REGION Network 5
   RUNG wire#powerrail
      { S7_Templates := "SrcType := Int" } EQ_Contact(in1 := #IN0, in2 := 2048)
      { S7_GenerateENO := "TRUE" } Move(in := 4, out1 => #OUT1)
   END_RUNG
   // the same network as SCL:
   IF #IN0 = 2048 THEN #OUT1 := 4; END_IF;
END_REGION

REGION Network 6
   RUNG wire#powerrail
      { S7_Templates := "SrcType := Int" } EQ_Contact(in1 := #IN0, in2 := 4096)
      { S7_GenerateENO := "TRUE" } Move(in := 5, out1 => #OUT1)
   END_RUNG
   // the same network as SCL:
   IF #IN0 = 4096 THEN #OUT1 := 5; END_IF;
END_REGION

REGION Network 7
   RUNG wire#powerrail
      { S7_Templates := "SrcType := Int" } EQ_Contact(in1 := #IN0, in2 := 8192)
      { S7_GenerateENO := "TRUE" } Move(in := 6, out1 => #OUT1)
   END_RUNG
   // the same network as SCL:
   IF #IN0 = 8192 THEN #OUT1 := 6; END_IF;
END_REGION

REGION Network 8
   RUNG wire#powerrail
      { S7_Templates := "SrcType := Int" } EQ_Contact(in1 := #IN0, in2 := 16384)
      { S7_GenerateENO := "TRUE" } Move(in := 7, out1 => #OUT1)
   END_RUNG
   // the same network as SCL:
   IF #IN0 = 16384 THEN #OUT1 := 7; END_IF;
END_REGION

REGION Network 9
   RUNG wire#powerrail
      { S7_Templates := "SrcType := Int" } EQ_Contact(in1 := #IN0, in2 := -32768)
      { S7_GenerateENO := "TRUE" } Move(in := 8, out1 => #OUT1)
   END_RUNG
   // the same network as SCL:
   IF #IN0 = (-32768) THEN #OUT1 := 8; END_IF;
END_REGION

REGION Network 10
   RUNG wire#powerrail
      { S7_Templates := "SrcType := Int" } EQ_Contact(in1 := #IN0, in2 := 1)
      { S7_GenerateENO := "TRUE" } Move(in := 9, out1 => #OUT1)
   END_RUNG
   // the same network as SCL:
   IF #IN0 = 1 THEN #OUT1 := 9; END_IF;
END_REGION

REGION Network 11
   RUNG wire#powerrail
      { S7_Templates := "SrcType := Int" } EQ_Contact(in1 := #IN0, in2 := 2)
      { S7_GenerateENO := "TRUE" } Move(in := 10, out1 => #OUT1)
   END_RUNG
   // the same network as SCL:
   IF #IN0 = 2 THEN #OUT1 := 10; END_IF;
END_REGION

REGION Network 12
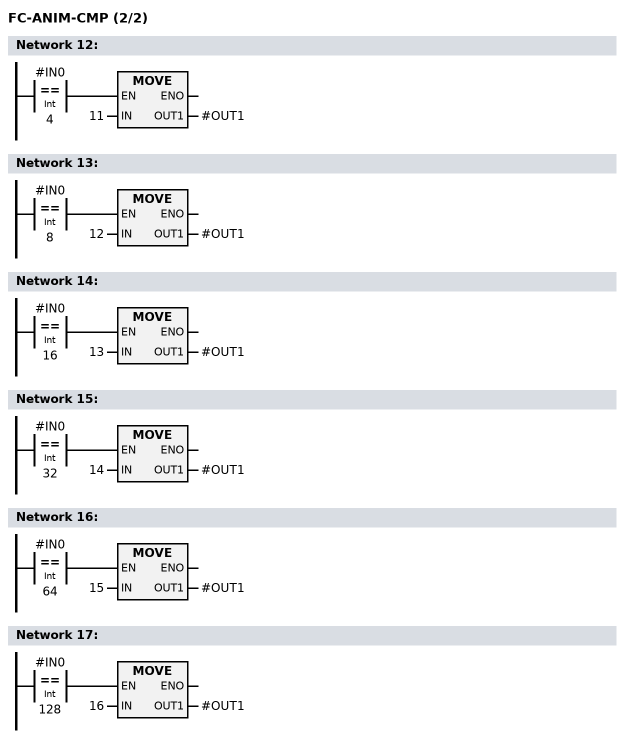
   RUNG wire#powerrail
      { S7_Templates := "SrcType := Int" } EQ_Contact(in1 := #IN0, in2 := 4)
      { S7_GenerateENO := "TRUE" } Move(in := 11, out1 => #OUT1)
   END_RUNG
   // the same network as SCL:
   IF #IN0 = 4 THEN #OUT1 := 11; END_IF;
END_REGION

REGION Network 13
   RUNG wire#powerrail
      { S7_Templates := "SrcType := Int" } EQ_Contact(in1 := #IN0, in2 := 8)
      { S7_GenerateENO := "TRUE" } Move(in := 12, out1 => #OUT1)
   END_RUNG
   // the same network as SCL:
   IF #IN0 = 8 THEN #OUT1 := 12; END_IF;
END_REGION

REGION Network 14
   RUNG wire#powerrail
      { S7_Templates := "SrcType := Int" } EQ_Contact(in1 := #IN0, in2 := 16)
      { S7_GenerateENO := "TRUE" } Move(in := 13, out1 => #OUT1)
   END_RUNG
   // the same network as SCL:
   IF #IN0 = 16 THEN #OUT1 := 13; END_IF;
END_REGION

REGION Network 15
   RUNG wire#powerrail
      { S7_Templates := "SrcType := Int" } EQ_Contact(in1 := #IN0, in2 := 32)
      { S7_GenerateENO := "TRUE" } Move(in := 14, out1 => #OUT1)
   END_RUNG
   // the same network as SCL:
   IF #IN0 = 32 THEN #OUT1 := 14; END_IF;
END_REGION

REGION Network 16
   RUNG wire#powerrail
      { S7_Templates := "SrcType := Int" } EQ_Contact(in1 := #IN0, in2 := 64)
      { S7_GenerateENO := "TRUE" } Move(in := 15, out1 => #OUT1)
   END_RUNG
   // the same network as SCL:
   IF #IN0 = 64 THEN #OUT1 := 15; END_IF;
END_REGION

REGION Network 17
   RUNG wire#powerrail
      { S7_Templates := "SrcType := Int" } EQ_Contact(in1 := #IN0, in2 := 128)
      { S7_GenerateENO := "TRUE" } Move(in := 16, out1 => #OUT1)
   END_RUNG
   // the same network as SCL:
   IF #IN0 = 128 THEN #OUT1 := 16; END_IF;
END_REGION
END_FUNCTION

// folder: Secadores/Alta

FUNCTION "EnclavSecAltaMTA" : Void   // FC12, LAD
{ S7_Optimized_Access := 'FALSE' }
VERSION : 0.1
BEGIN

REGION Network 1: Arranque automático MS050
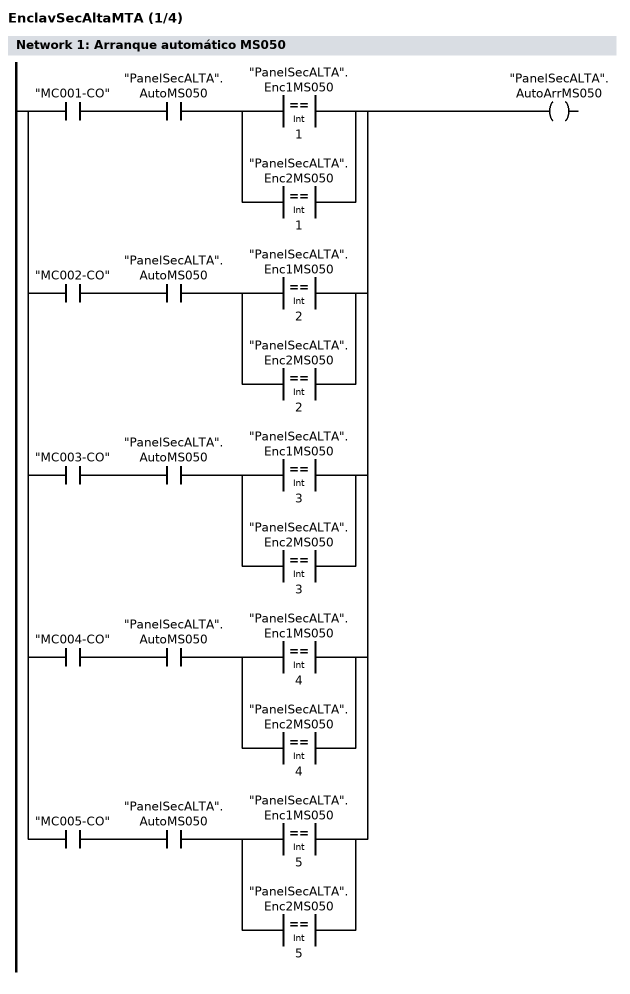
   "PanelSecALTA".AutoArrMS050 := ("MC001-CO" AND "PanelSecALTA".AutoMS050 AND (("PanelSecALTA".Enc1MS050 = 1) OR ("PanelSecALTA".Enc2MS050 = 1))) OR ("MC002-CO" AND "PanelSecALTA".AutoMS050 AND (("PanelSecALTA".Enc1MS050 = 2) OR ("PanelSecALTA".Enc2MS050 = 2))) OR ("MC003-CO" AND "PanelSecALTA".AutoMS050 AND (("PanelSecALTA".Enc1MS050 = 3) OR ("PanelSecALTA".Enc2MS050 = 3))) OR ("MC004-CO" AND "PanelSecALTA".AutoMS050 AND (("PanelSecALTA".Enc1MS050 = 4) OR ("PanelSecALTA".Enc2MS050 = 4))) OR ("MC005-CO" AND "PanelSecALTA".AutoMS050 AND (("PanelSecALTA".Enc1MS050 = 5) OR ("PanelSecALTA".Enc2MS050 = 5)));
END_REGION

REGION Network 2: Arranque automático MS051
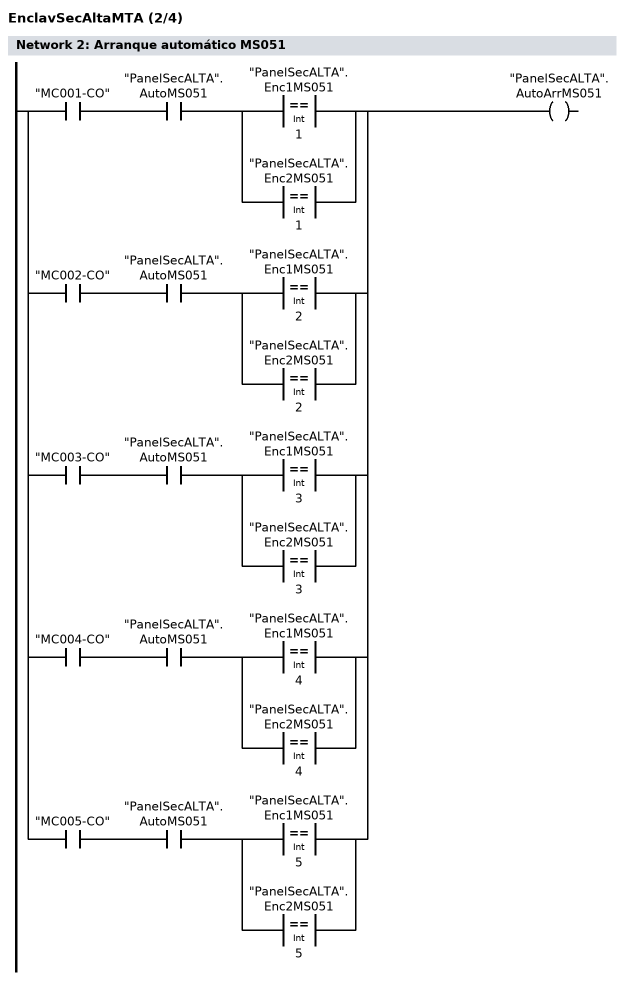
   "PanelSecALTA".AutoArrMS051 := ("MC001-CO" AND "PanelSecALTA".AutoMS051 AND (("PanelSecALTA".Enc1MS051 = 1) OR ("PanelSecALTA".Enc2MS051 = 1))) OR ("MC002-CO" AND "PanelSecALTA".AutoMS051 AND (("PanelSecALTA".Enc1MS051 = 2) OR ("PanelSecALTA".Enc2MS051 = 2))) OR ("MC003-CO" AND "PanelSecALTA".AutoMS051 AND (("PanelSecALTA".Enc1MS051 = 3) OR ("PanelSecALTA".Enc2MS051 = 3))) OR ("MC004-CO" AND "PanelSecALTA".AutoMS051 AND (("PanelSecALTA".Enc1MS051 = 4) OR ("PanelSecALTA".Enc2MS051 = 4))) OR ("MC005-CO" AND "PanelSecALTA".AutoMS051 AND (("PanelSecALTA".Enc1MS051 = 5) OR ("PanelSecALTA".Enc2MS051 = 5)));
END_REGION

REGION Network 3: Arranque automático MS052
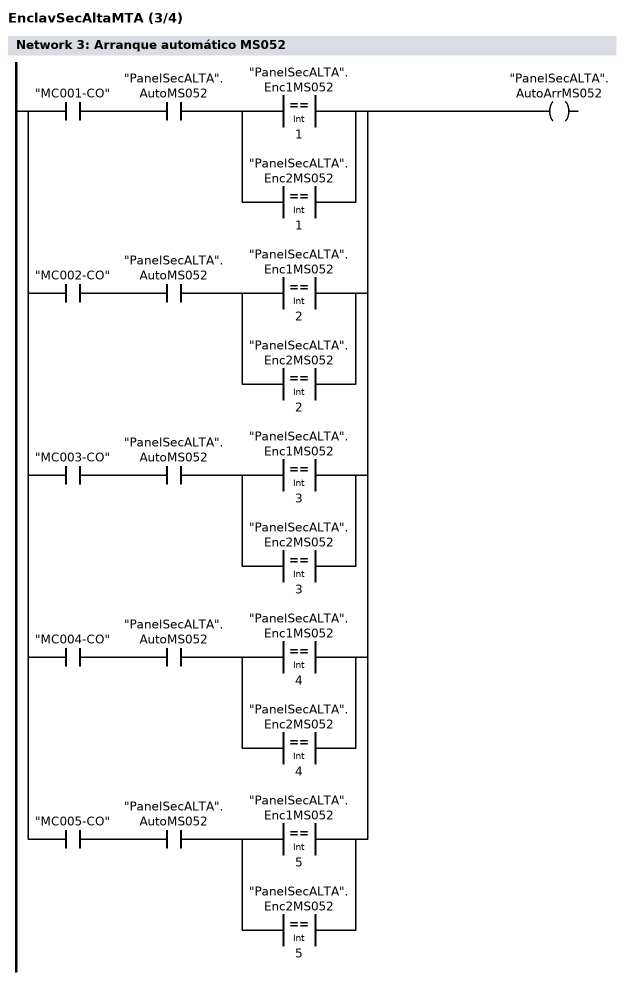
   "PanelSecALTA".AutoArrMS052 := ("MC001-CO" AND "PanelSecALTA".AutoMS052 AND (("PanelSecALTA".Enc1MS052 = 1) OR ("PanelSecALTA".Enc2MS052 = 1))) OR ("MC002-CO" AND "PanelSecALTA".AutoMS052 AND (("PanelSecALTA".Enc1MS052 = 2) OR ("PanelSecALTA".Enc2MS052 = 2))) OR ("MC003-CO" AND "PanelSecALTA".AutoMS052 AND (("PanelSecALTA".Enc1MS052 = 3) OR ("PanelSecALTA".Enc2MS052 = 3))) OR ("MC004-CO" AND "PanelSecALTA".AutoMS052 AND (("PanelSecALTA".Enc1MS052 = 4) OR ("PanelSecALTA".Enc2MS052 = 4))) OR ("MC005-CO" AND "PanelSecALTA".AutoMS052 AND (("PanelSecALTA".Enc1MS052 = 5) OR ("PanelSecALTA".Enc2MS052 = 5)));
END_REGION

REGION Network 4: Arranque automático MS053
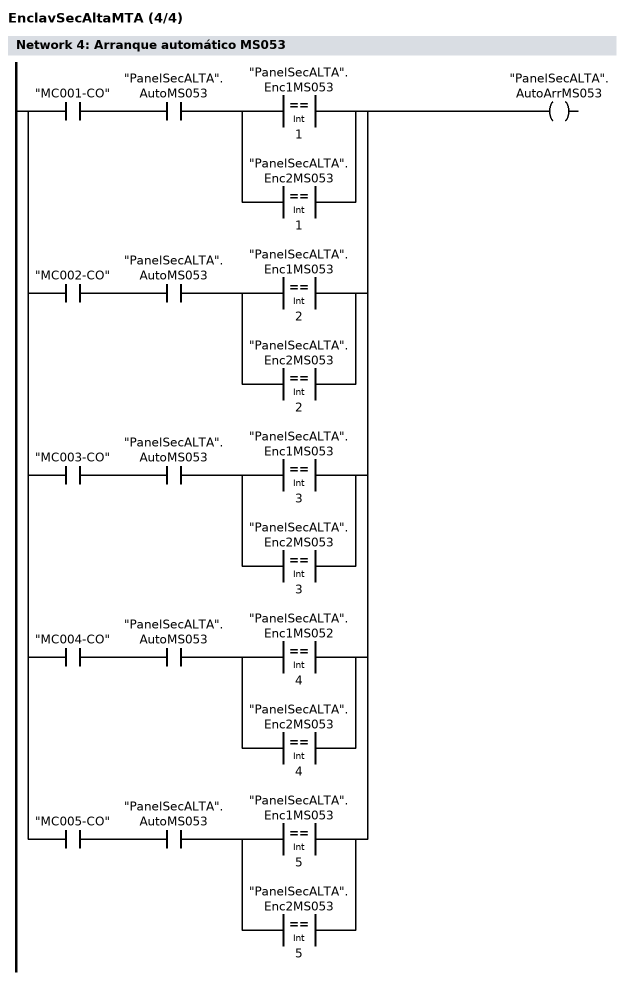
   "PanelSecALTA".AutoArrMS053 := ("MC001-CO" AND "PanelSecALTA".AutoMS053 AND (("PanelSecALTA".Enc1MS053 = 1) OR ("PanelSecALTA".Enc2MS053 = 1))) OR ("MC002-CO" AND "PanelSecALTA".AutoMS053 AND (("PanelSecALTA".Enc1MS053 = 2) OR ("PanelSecALTA".Enc2MS053 = 2))) OR ("MC003-CO" AND "PanelSecALTA".AutoMS053 AND (("PanelSecALTA".Enc1MS053 = 3) OR ("PanelSecALTA".Enc2MS053 = 3))) OR ("MC004-CO" AND "PanelSecALTA".AutoMS053 AND (("PanelSecALTA".Enc1MS052 = 4) OR ("PanelSecALTA".Enc2MS053 = 4))) OR ("MC005-CO" AND "PanelSecALTA".AutoMS053 AND (("PanelSecALTA".Enc1MS053 = 5) OR ("PanelSecALTA".Enc2MS053 = 5)));
END_REGION
END_FUNCTION

// folder: Torres de Agua/Torres Cavaleto

FUNCTION "TorresCavaletoMTA" : Void   // FC14, LAD
{ S7_Optimized_Access := 'FALSE' }
VERSION : 0.1
BEGIN

REGION Network 1: Comandos MV030 / Comandos desde Panel para MV030 - Ventilador 2 Torres de enfriamiento Cavaleto
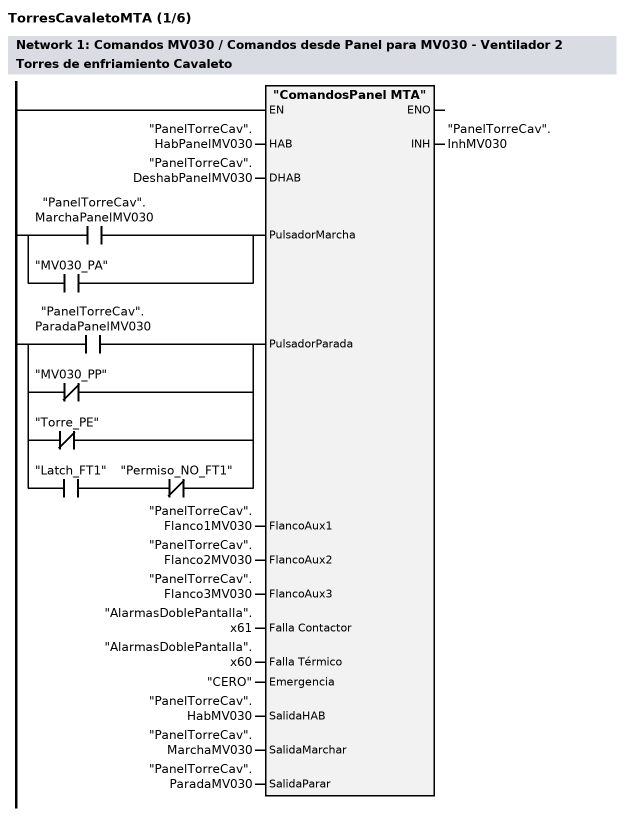
   RUNG wire#powerrail
      "ComandosPanel MTA"(PulsadorMarcha := wire#w1, PulsadorParada := wire#w2, HAB := "PanelTorreCav".HabPanelMV030, DHAB := "PanelTorreCav".DeshabPanelMV030, FlancoAux1 := "PanelTorreCav".Flanco1MV030, FlancoAux2 := "PanelTorreCav".Flanco2MV030, FlancoAux3 := "PanelTorreCav".Flanco3MV030, "Falla Contactor" := "AlarmasDoblePantalla".x61, "Falla Térmico" := "AlarmasDoblePantalla".x60, Emergencia := "CERO", SalidaHAB := "PanelTorreCav".HabMV030, SalidaMarchar := "PanelTorreCav".MarchaMV030, SalidaParar := "PanelTorreCav".ParadaMV030, INH => "PanelTorreCav".InhMV030)
   END_RUNG
   RUNG wire#powerrail
      Contact( "PanelTorreCav".MarchaPanelMV030 )
   END_RUNG wire#w1
   RUNG wire#powerrail
      Contact( "MV030_PA" )
   END_RUNG wire#w1
   RUNG wire#powerrail
      Contact( "PanelTorreCav".ParadaPanelMV030 )
   END_RUNG wire#w2
   RUNG wire#powerrail
      I_Contact( "MV030_PP" )
   END_RUNG wire#w2
   RUNG wire#powerrail
      I_Contact( "Torre_PE" )
   END_RUNG wire#w2
   RUNG wire#powerrail
      Contact( "Latch_FT1" )
      I_Contact( "Permiso_NO_FT1" )
   END_RUNG wire#w2
   // the same network as SCL:
   "ComandosPanel MTA"(HAB := "PanelTorreCav".HabPanelMV030,
                       DHAB := "PanelTorreCav".DeshabPanelMV030,
                       PulsadorMarcha := "PanelTorreCav".MarchaPanelMV030 OR "MV030_PA",
                       PulsadorParada := "PanelTorreCav".ParadaPanelMV030 OR NOT "MV030_PP" OR NOT "Torre_PE" OR ("Latch_FT1" AND NOT "Permiso_NO_FT1"),
                       FlancoAux1 := "PanelTorreCav".Flanco1MV030,
                       FlancoAux2 := "PanelTorreCav".Flanco2MV030,
                       FlancoAux3 := "PanelTorreCav".Flanco3MV030,
                       "Falla Contactor" := "AlarmasDoblePantalla".x61,
                       "Falla Térmico" := "AlarmasDoblePantalla".x60,
                       Emergencia := "CERO",
                       SalidaHAB := "PanelTorreCav".HabMV030,
                       SalidaMarchar := "PanelTorreCav".MarchaMV030,
                       SalidaParar := "PanelTorreCav".ParadaMV030,
                       INH => "PanelTorreCav".InhMV030);
END_REGION

REGION Network 2: Comandos MV031 / Comandos desde Panel para MV031 - Ventilador 1 Torres de enfriamiento Cavaleto
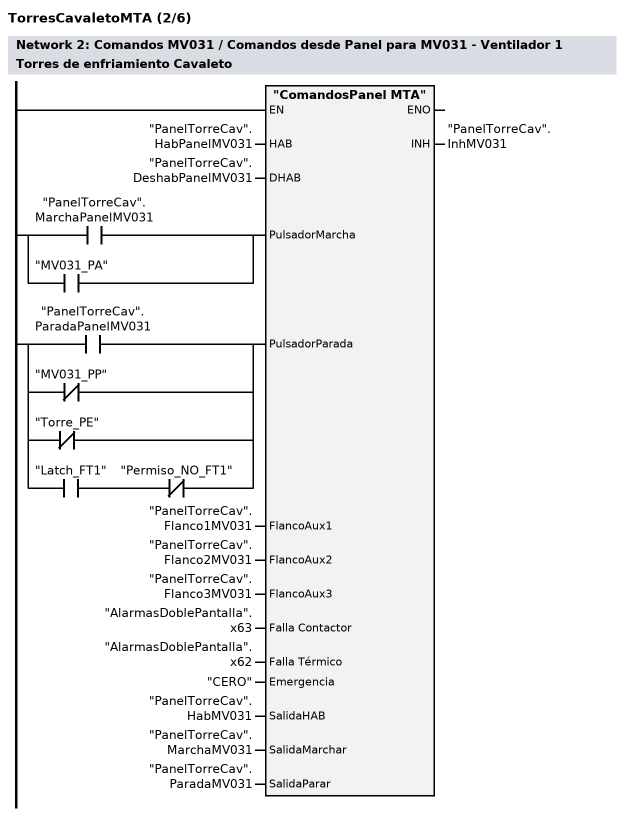
   RUNG wire#powerrail
      "ComandosPanel MTA"(PulsadorMarcha := wire#w1, PulsadorParada := wire#w2, HAB := "PanelTorreCav".HabPanelMV031, DHAB := "PanelTorreCav".DeshabPanelMV031, FlancoAux1 := "PanelTorreCav".Flanco1MV031, FlancoAux2 := "PanelTorreCav".Flanco2MV031, FlancoAux3 := "PanelTorreCav".Flanco3MV031, "Falla Contactor" := "AlarmasDoblePantalla".x63, "Falla Térmico" := "AlarmasDoblePantalla".x62, Emergencia := "CERO", SalidaHAB := "PanelTorreCav".HabMV031, SalidaMarchar := "PanelTorreCav".MarchaMV031, SalidaParar := "PanelTorreCav".ParadaMV031, INH => "PanelTorreCav".InhMV031)
   END_RUNG
   RUNG wire#powerrail
      Contact( "PanelTorreCav".MarchaPanelMV031 )
   END_RUNG wire#w1
   RUNG wire#powerrail
      Contact( "MV031_PA" )
   END_RUNG wire#w1
   RUNG wire#powerrail
      Contact( "PanelTorreCav".ParadaPanelMV031 )
   END_RUNG wire#w2
   RUNG wire#powerrail
      I_Contact( "MV031_PP" )
   END_RUNG wire#w2
   RUNG wire#powerrail
      I_Contact( "Torre_PE" )
   END_RUNG wire#w2
   RUNG wire#powerrail
      Contact( "Latch_FT1" )
      I_Contact( "Permiso_NO_FT1" )
   END_RUNG wire#w2
   // the same network as SCL:
   "ComandosPanel MTA"(HAB := "PanelTorreCav".HabPanelMV031,
                       DHAB := "PanelTorreCav".DeshabPanelMV031,
                       PulsadorMarcha := "PanelTorreCav".MarchaPanelMV031 OR "MV031_PA",
                       PulsadorParada := "PanelTorreCav".ParadaPanelMV031 OR NOT "MV031_PP" OR NOT "Torre_PE" OR ("Latch_FT1" AND NOT "Permiso_NO_FT1"),
                       FlancoAux1 := "PanelTorreCav".Flanco1MV031,
                       FlancoAux2 := "PanelTorreCav".Flanco2MV031,
                       FlancoAux3 := "PanelTorreCav".Flanco3MV031,
                       "Falla Contactor" := "AlarmasDoblePantalla".x63,
                       "Falla Térmico" := "AlarmasDoblePantalla".x62,
                       Emergencia := "CERO",
                       SalidaHAB := "PanelTorreCav".HabMV031,
                       SalidaMarchar := "PanelTorreCav".MarchaMV031,
                       SalidaParar := "PanelTorreCav".ParadaMV031,
                       INH => "PanelTorreCav".InhMV031);
END_REGION

REGION Network 3: Comandos MP014 / Comandos desde Panel para P014 - Bomba 1 Torres de enfriamiento Cavaleto
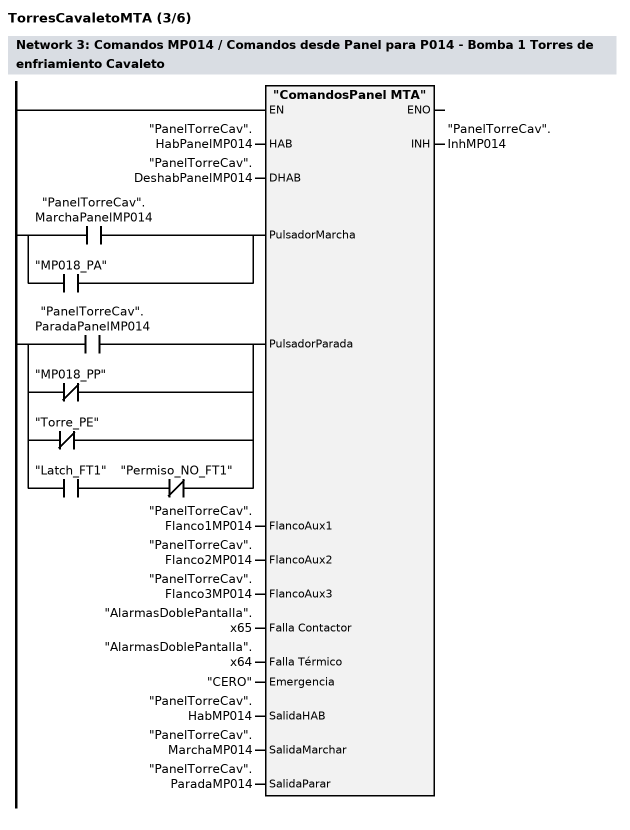
   RUNG wire#powerrail
      "ComandosPanel MTA"(PulsadorMarcha := wire#w1, PulsadorParada := wire#w2, HAB := "PanelTorreCav".HabPanelMP014, DHAB := "PanelTorreCav".DeshabPanelMP014, FlancoAux1 := "PanelTorreCav".Flanco1MP014, FlancoAux2 := "PanelTorreCav".Flanco2MP014, FlancoAux3 := "PanelTorreCav".Flanco3MP014, "Falla Contactor" := "AlarmasDoblePantalla".x65, "Falla Térmico" := "AlarmasDoblePantalla".x64, Emergencia := "CERO", SalidaHAB := "PanelTorreCav".HabMP014, SalidaMarchar := "PanelTorreCav".MarchaMP014, SalidaParar := "PanelTorreCav".ParadaMP014, INH => "PanelTorreCav".InhMP014)
   END_RUNG
   RUNG wire#powerrail
      Contact( "PanelTorreCav".MarchaPanelMP014 )
   END_RUNG wire#w1
   RUNG wire#powerrail
      Contact( "MP018_PA" )
   END_RUNG wire#w1
   RUNG wire#powerrail
      Contact( "PanelTorreCav".ParadaPanelMP014 )
   END_RUNG wire#w2
   RUNG wire#powerrail
      I_Contact( "MP018_PP" )
   END_RUNG wire#w2
   RUNG wire#powerrail
      I_Contact( "Torre_PE" )
   END_RUNG wire#w2
   RUNG wire#powerrail
      Contact( "Latch_FT1" )
      I_Contact( "Permiso_NO_FT1" )
   END_RUNG wire#w2
   // the same network as SCL:
   "ComandosPanel MTA"(HAB := "PanelTorreCav".HabPanelMP014,
                       DHAB := "PanelTorreCav".DeshabPanelMP014,
                       PulsadorMarcha := "PanelTorreCav".MarchaPanelMP014 OR "MP018_PA",
                       PulsadorParada := "PanelTorreCav".ParadaPanelMP014 OR NOT "MP018_PP" OR NOT "Torre_PE" OR ("Latch_FT1" AND NOT "Permiso_NO_FT1"),
                       FlancoAux1 := "PanelTorreCav".Flanco1MP014,
                       FlancoAux2 := "PanelTorreCav".Flanco2MP014,
                       FlancoAux3 := "PanelTorreCav".Flanco3MP014,
                       "Falla Contactor" := "AlarmasDoblePantalla".x65,
                       "Falla Térmico" := "AlarmasDoblePantalla".x64,
                       Emergencia := "CERO",
                       SalidaHAB := "PanelTorreCav".HabMP014,
                       SalidaMarchar := "PanelTorreCav".MarchaMP014,
                       SalidaParar := "PanelTorreCav".ParadaMP014,
                       INH => "PanelTorreCav".InhMP014);
END_REGION

REGION Network 4: Comandos MP015 / Comandos desde Panel para P015 - Bomba 2 Torres de enfriamiento Cavaleto
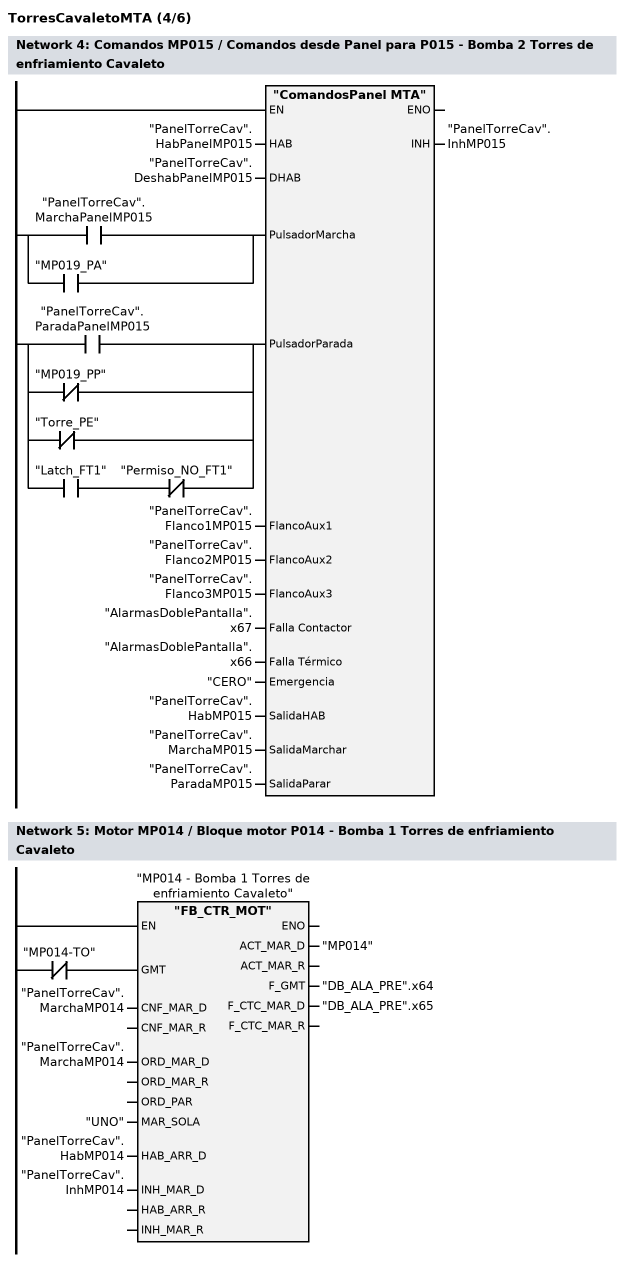
   RUNG wire#powerrail
      "ComandosPanel MTA"(PulsadorMarcha := wire#w1, PulsadorParada := wire#w2, HAB := "PanelTorreCav".HabPanelMP015, DHAB := "PanelTorreCav".DeshabPanelMP015, FlancoAux1 := "PanelTorreCav".Flanco1MP015, FlancoAux2 := "PanelTorreCav".Flanco2MP015, FlancoAux3 := "PanelTorreCav".Flanco3MP015, "Falla Contactor" := "AlarmasDoblePantalla".x67, "Falla Térmico" := "AlarmasDoblePantalla".x66, Emergencia := "CERO", SalidaHAB := "PanelTorreCav".HabMP015, SalidaMarchar := "PanelTorreCav".MarchaMP015, SalidaParar := "PanelTorreCav".ParadaMP015, INH => "PanelTorreCav".InhMP015)
   END_RUNG
   RUNG wire#powerrail
      Contact( "PanelTorreCav".MarchaPanelMP015 )
   END_RUNG wire#w1
   RUNG wire#powerrail
      Contact( "MP019_PA" )
   END_RUNG wire#w1
   RUNG wire#powerrail
      Contact( "PanelTorreCav".ParadaPanelMP015 )
   END_RUNG wire#w2
   RUNG wire#powerrail
      I_Contact( "MP019_PP" )
   END_RUNG wire#w2
   RUNG wire#powerrail
      I_Contact( "Torre_PE" )
   END_RUNG wire#w2
   RUNG wire#powerrail
      Contact( "Latch_FT1" )
      I_Contact( "Permiso_NO_FT1" )
   END_RUNG wire#w2
   // the same network as SCL:
   "ComandosPanel MTA"(HAB := "PanelTorreCav".HabPanelMP015,
                       DHAB := "PanelTorreCav".DeshabPanelMP015,
                       PulsadorMarcha := "PanelTorreCav".MarchaPanelMP015 OR "MP019_PA",
                       PulsadorParada := "PanelTorreCav".ParadaPanelMP015 OR NOT "MP019_PP" OR NOT "Torre_PE" OR ("Latch_FT1" AND NOT "Permiso_NO_FT1"),
                       FlancoAux1 := "PanelTorreCav".Flanco1MP015,
                       FlancoAux2 := "PanelTorreCav".Flanco2MP015,
                       FlancoAux3 := "PanelTorreCav".Flanco3MP015,
                       "Falla Contactor" := "AlarmasDoblePantalla".x67,
                       "Falla Térmico" := "AlarmasDoblePantalla".x66,
                       Emergencia := "CERO",
                       SalidaHAB := "PanelTorreCav".HabMP015,
                       SalidaMarchar := "PanelTorreCav".MarchaMP015,
                       SalidaParar := "PanelTorreCav".ParadaMP015,
                       INH => "PanelTorreCav".InhMP015);
END_REGION

REGION Network 5: Motor MP014 / Bloque motor P014 - Bomba 1 Torres de enfriamiento Cavaleto
   RUNG wire#powerrail
      "MP014 - Bomba 1 Torres de enfriamiento Cavaleto"(CNF_MAR_D := "PanelTorreCav".MarchaMP014, CNF_MAR_R :=, ORD_MAR_D := "PanelTorreCav".MarchaMP014, ORD_MAR_R :=, ORD_PAR :=, MAR_SOLA := "UNO", HAB_ARR_D := "PanelTorreCav".HabMP014, INH_MAR_D := "PanelTorreCav".InhMP014, HAB_ARR_R :=, INH_MAR_R :=, ACT_MAR_D => "MP014", ACT_MAR_R =>, F_GMT => "DB_ALA_PRE".x64, F_CTC_MAR_D => "DB_ALA_PRE".x65, F_CTC_MAR_R =>, GMT := wire#w1)
   END_RUNG
   RUNG wire#powerrail
      I_Contact( "MP014-TO" )
   END_RUNG wire#w1
   // the same network as SCL:
   "MP014 - Bomba 1 Torres de enfriamiento Cavaleto"(GMT := NOT "MP014-TO",   // "FB_CTR_MOT"
                           CNF_MAR_D := "PanelTorreCav".MarchaMP014,
                           ORD_MAR_D := "PanelTorreCav".MarchaMP014,
                           MAR_SOLA := "UNO",
                           HAB_ARR_D := "PanelTorreCav".HabMP014,
                           INH_MAR_D := "PanelTorreCav".InhMP014,
                           ACT_MAR_D => "MP014",
                           F_GMT => "DB_ALA_PRE".x64,
                           F_CTC_MAR_D => "DB_ALA_PRE".x65);
END_REGION

REGION Network 6: Motor MP015 / Bloque motor P015 - Bomba 2 Torres de enfriamiento Cavaleto
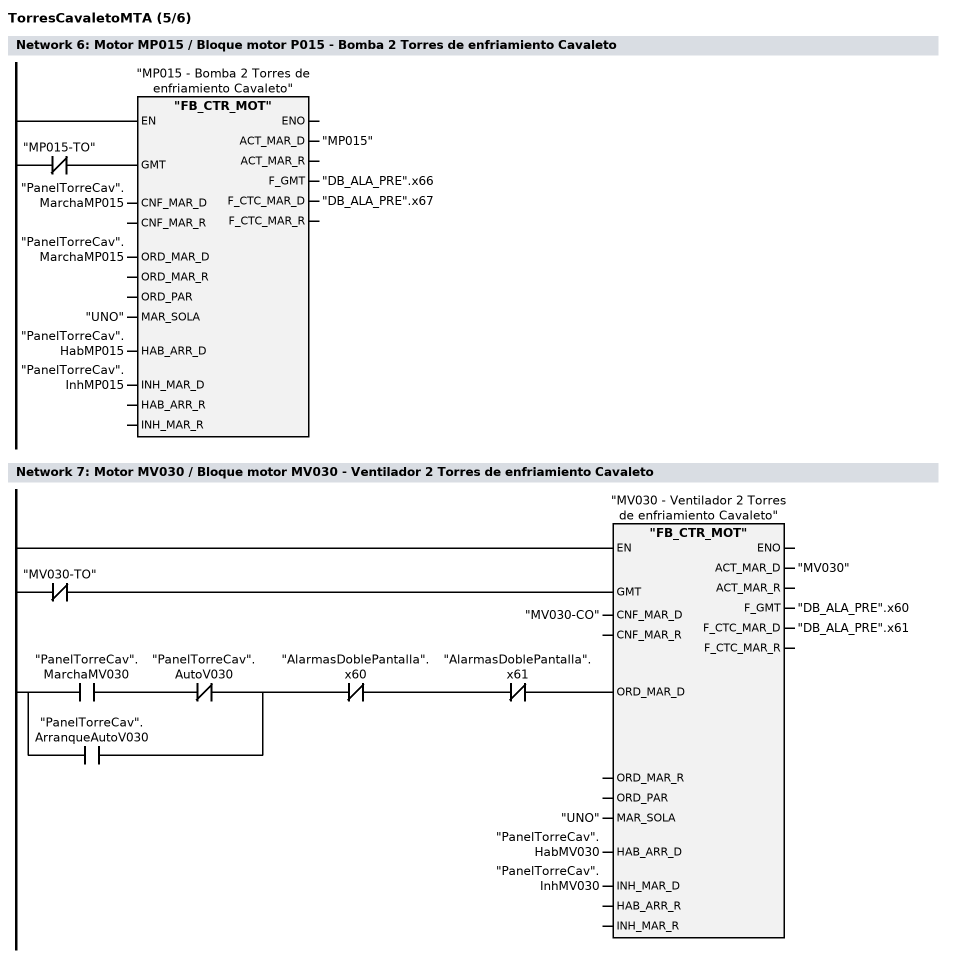
   RUNG wire#powerrail
      "MP015 - Bomba 2 Torres de enfriamiento Cavaleto"(CNF_MAR_D := "PanelTorreCav".MarchaMP015, CNF_MAR_R :=, ORD_MAR_D := "PanelTorreCav".MarchaMP015, ORD_MAR_R :=, ORD_PAR :=, MAR_SOLA := "UNO", HAB_ARR_D := "PanelTorreCav".HabMP015, INH_MAR_D := "PanelTorreCav".InhMP015, HAB_ARR_R :=, INH_MAR_R :=, ACT_MAR_D => "MP015", ACT_MAR_R =>, F_GMT => "DB_ALA_PRE".x66, F_CTC_MAR_D => "DB_ALA_PRE".x67, F_CTC_MAR_R =>, GMT := wire#w1)
   END_RUNG
   RUNG wire#powerrail
      I_Contact( "MP015-TO" )
   END_RUNG wire#w1
   // the same network as SCL:
   "MP015 - Bomba 2 Torres de enfriamiento Cavaleto"(GMT := NOT "MP015-TO",   // "FB_CTR_MOT"
                           CNF_MAR_D := "PanelTorreCav".MarchaMP015,
                           ORD_MAR_D := "PanelTorreCav".MarchaMP015,
                           MAR_SOLA := "UNO",
                           HAB_ARR_D := "PanelTorreCav".HabMP015,
                           INH_MAR_D := "PanelTorreCav".InhMP015,
                           ACT_MAR_D => "MP015",
                           F_GMT => "DB_ALA_PRE".x66,
                           F_CTC_MAR_D => "DB_ALA_PRE".x67);
END_REGION

REGION Network 7: Motor MV030 / Bloque motor MV030 - Ventilador 2 Torres de enfriamiento Cavaleto
   RUNG wire#powerrail
      "MV030 - Ventilador 2 Torres de enfriamiento Cavaleto"(GMT := wire#w1, ORD_MAR_D := wire#w3, CNF_MAR_D := "MV030-CO", CNF_MAR_R :=, ORD_MAR_R :=, ORD_PAR :=, MAR_SOLA := "UNO", HAB_ARR_D := "PanelTorreCav".HabMV030, INH_MAR_D := "PanelTorreCav".InhMV030, HAB_ARR_R :=, INH_MAR_R :=, ACT_MAR_D => "MV030", ACT_MAR_R =>, F_GMT => "DB_ALA_PRE".x60, F_CTC_MAR_D => "DB_ALA_PRE".x61, F_CTC_MAR_R =>)
   END_RUNG
   RUNG wire#powerrail
      I_Contact( "MV030-TO" )
   END_RUNG wire#w1
   RUNG wire#powerrail
      Contact( "PanelTorreCav".MarchaMV030 )
      I_Contact( "PanelTorreCav".AutoV030 )
      wire#w2
      I_Contact( "AlarmasDoblePantalla".x60 )
      I_Contact( "AlarmasDoblePantalla".x61 )
   END_RUNG wire#w3
   RUNG wire#powerrail
      Contact( "PanelTorreCav".ArranqueAutoV030 )
   END_RUNG wire#w2
   // the same network as SCL:
   "MV030 - Ventilador 2 Torres de enfriamiento Cavaleto"(GMT := NOT "MV030-TO",   // "FB_CTR_MOT"
                           CNF_MAR_D := "MV030-CO",
                           ORD_MAR_D := (("PanelTorreCav".MarchaMV030 AND NOT "PanelTorreCav".AutoV030) OR "PanelTorreCav".ArranqueAutoV030) AND NOT "AlarmasDoblePantalla".x60 AND NOT "AlarmasDoblePantalla".x61,
                           MAR_SOLA := "UNO",
                           HAB_ARR_D := "PanelTorreCav".HabMV030,
                           INH_MAR_D := "PanelTorreCav".InhMV030,
                           ACT_MAR_D => "MV030",
                           F_GMT => "DB_ALA_PRE".x60,
                           F_CTC_MAR_D => "DB_ALA_PRE".x61);
END_REGION

REGION Network 8: Motor MV031 / Bloque motorMV031 - Ventilador 1 Torres de enfriamiento Cavaleto
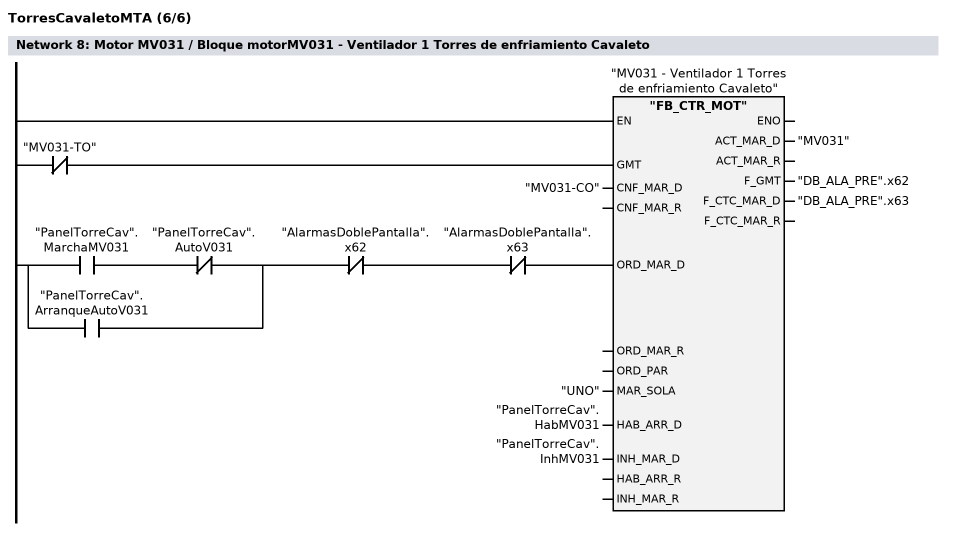
   RUNG wire#powerrail
      "MV031 - Ventilador 1 Torres de enfriamiento Cavaleto"(GMT := wire#w1, ORD_MAR_D := wire#w3, CNF_MAR_D := "MV031-CO", CNF_MAR_R :=, ORD_MAR_R :=, ORD_PAR :=, MAR_SOLA := "UNO", HAB_ARR_D := "PanelTorreCav".HabMV031, INH_MAR_D := "PanelTorreCav".InhMV031, HAB_ARR_R :=, INH_MAR_R :=, ACT_MAR_D => "MV031", ACT_MAR_R =>, F_GMT => "DB_ALA_PRE".x62, F_CTC_MAR_D => "DB_ALA_PRE".x63, F_CTC_MAR_R =>)
   END_RUNG
   RUNG wire#powerrail
      I_Contact( "MV031-TO" )
   END_RUNG wire#w1
   RUNG wire#powerrail
      Contact( "PanelTorreCav".MarchaMV031 )
      I_Contact( "PanelTorreCav".AutoV031 )
      wire#w2
      I_Contact( "AlarmasDoblePantalla".x62 )
      I_Contact( "AlarmasDoblePantalla".x63 )
   END_RUNG wire#w3
   RUNG wire#powerrail
      Contact( "PanelTorreCav".ArranqueAutoV031 )
   END_RUNG wire#w2
   // the same network as SCL:
   "MV031 - Ventilador 1 Torres de enfriamiento Cavaleto"(GMT := NOT "MV031-TO",   // "FB_CTR_MOT"
                           CNF_MAR_D := "MV031-CO",
                           ORD_MAR_D := (("PanelTorreCav".MarchaMV031 AND NOT "PanelTorreCav".AutoV031) OR "PanelTorreCav".ArranqueAutoV031) AND NOT "AlarmasDoblePantalla".x62 AND NOT "AlarmasDoblePantalla".x63,
                           MAR_SOLA := "UNO",
                           HAB_ARR_D := "PanelTorreCav".HabMV031,
                           INH_MAR_D := "PanelTorreCav".InhMV031,
                           ACT_MAR_D => "MV031",
                           F_GMT => "DB_ALA_PRE".x62,
                           F_CTC_MAR_D => "DB_ALA_PRE".x63);
END_REGION
END_FUNCTION

// folder: Torres de Agua/Torres Chillers

FUNCTION "TorresAutoMTA" : Void   // FC9, LAD
{ S7_Optimized_Access := 'FALSE' }
VERSION : 0.1
BEGIN

REGION Network 1: Lectura Temperatura de Torres Chillers
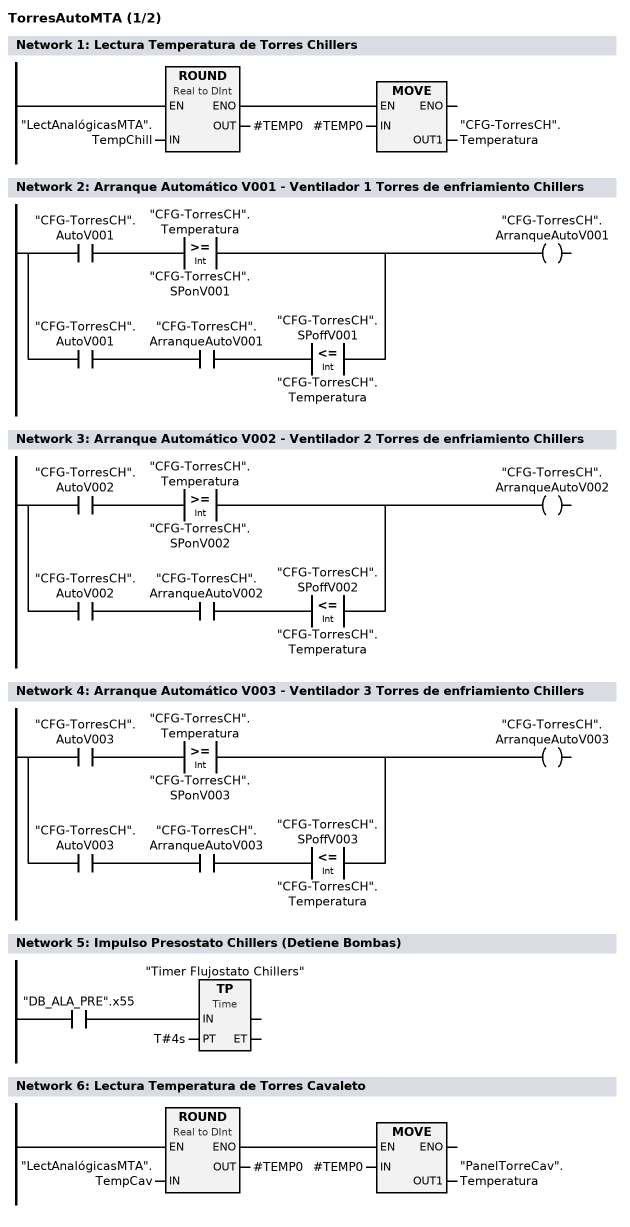
   RUNG wire#powerrail
      { S7_Templates := "[SrcType := Real, DestType := DInt]"; S7_GenerateENO := "TRUE" } Round(in := "LectAnalógicasMTA".TempChill, out => #TEMP0)
      { S7_GenerateENO := "TRUE" } Move(in := #TEMP0, out1 => "CFG-TorresCH".Temperatura)
   END_RUNG
   // the same network as SCL:
   // ENO of a box is taken as its EN; it also drops when the box reports an error
   #TEMP0 := ROUND("LectAnalógicasMTA".TempChill);
   "CFG-TorresCH".Temperatura := #TEMP0;
END_REGION

REGION Network 2: Arranque Automático V001 - Ventilador 1 Torres de enfriamiento Chillers
   "CFG-TorresCH".ArranqueAutoV001 := ("CFG-TorresCH".AutoV001 AND ("CFG-TorresCH".Temperatura >= "CFG-TorresCH".SPonV001)) OR ("CFG-TorresCH".AutoV001 AND "CFG-TorresCH".ArranqueAutoV001 AND ("CFG-TorresCH".SPoffV001 <= "CFG-TorresCH".Temperatura));
END_REGION

REGION Network 3: Arranque Automático V002 - Ventilador 2 Torres de enfriamiento Chillers
   "CFG-TorresCH".ArranqueAutoV002 := ("CFG-TorresCH".AutoV002 AND ("CFG-TorresCH".Temperatura >= "CFG-TorresCH".SPonV002)) OR ("CFG-TorresCH".AutoV002 AND "CFG-TorresCH".ArranqueAutoV002 AND ("CFG-TorresCH".SPoffV002 <= "CFG-TorresCH".Temperatura));
END_REGION

REGION Network 4: Arranque Automático V003 - Ventilador 3 Torres de enfriamiento Chillers
   "CFG-TorresCH".ArranqueAutoV003 := ("CFG-TorresCH".AutoV003 AND ("CFG-TorresCH".Temperatura >= "CFG-TorresCH".SPonV003)) OR ("CFG-TorresCH".AutoV003 AND "CFG-TorresCH".ArranqueAutoV003 AND ("CFG-TorresCH".SPoffV003 <= "CFG-TorresCH".Temperatura));
END_REGION

REGION Network 5: Impulso Presostato Chillers (Detiene Bombas)
   "Timer Flujostato Chillers".TP(in := "DB_ALA_PRE".x55, pt := T#4s);
END_REGION

REGION Network 6: Lectura Temperatura de Torres Cavaleto
   RUNG wire#powerrail
      { S7_Templates := "[SrcType := Real, DestType := DInt]"; S7_GenerateENO := "TRUE" } Round(in := "LectAnalógicasMTA".TempCav, out => #TEMP0)
      { S7_GenerateENO := "TRUE" } Move(in := #TEMP0, out1 => "PanelTorreCav".Temperatura)
   END_RUNG
   // the same network as SCL:
   // ENO of a box is taken as its EN; it also drops when the box reports an error
   #TEMP0 := ROUND("LectAnalógicasMTA".TempCav);
   "PanelTorreCav".Temperatura := #TEMP0;
END_REGION

REGION Network 7: Arranque Automático MV030 - Ventilador 1 Torres de enfriamiento Cavaleto
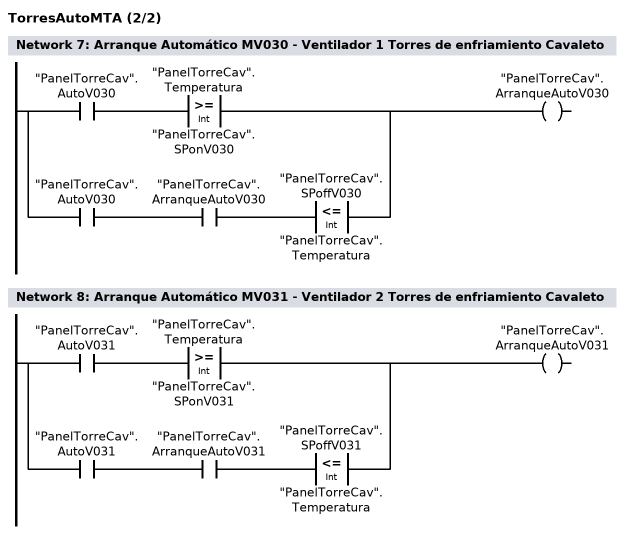
   "PanelTorreCav".ArranqueAutoV030 := ("PanelTorreCav".AutoV030 AND ("PanelTorreCav".Temperatura >= "PanelTorreCav".SPonV030)) OR ("PanelTorreCav".AutoV030 AND "PanelTorreCav".ArranqueAutoV030 AND ("PanelTorreCav".SPoffV030 <= "PanelTorreCav".Temperatura));
END_REGION

REGION Network 8: Arranque Automático MV031 - Ventilador 2 Torres de enfriamiento Cavaleto
   "PanelTorreCav".ArranqueAutoV031 := ("PanelTorreCav".AutoV031 AND ("PanelTorreCav".Temperatura >= "PanelTorreCav".SPonV031)) OR ("PanelTorreCav".AutoV031 AND "PanelTorreCav".ArranqueAutoV031 AND ("PanelTorreCav".SPoffV031 <= "PanelTorreCav".Temperatura));
END_REGION
END_FUNCTION

(* ===== HMI "HMI_RT_3" =====
connection "Conexión2-PLC_1": ETHERNET, SIMATIC S7 300/400 MPI
